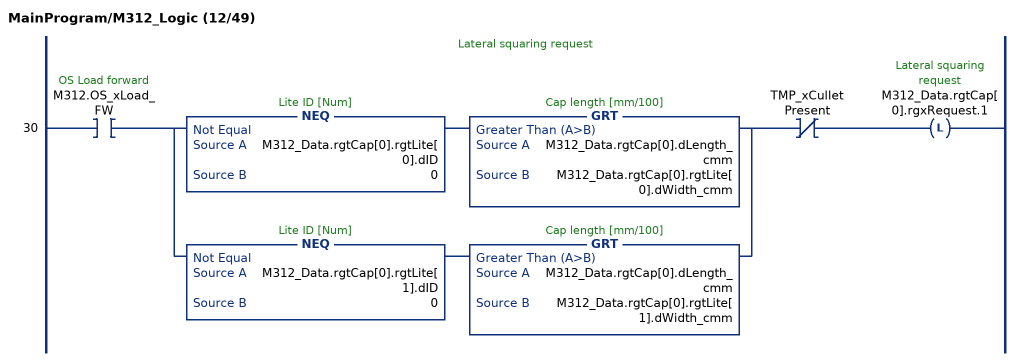
   // Lateral squaring request
   30: XIC(M312.OS_xLoad_FW)[NEQ(M312_Data.rgtCap[0].rgtLite[0].dID,0) GRT(M312_Data.rgtCap[0].dLength_cmm,M312_Data.rgtCap[0].rgtLite[0].dWidth_cmm) ,NEQ(M312_Data.rgtCap[0].rgtLite[1].dID,0) GRT(M312_Data.rgtCap[0].dLength_cmm,M312_Data.rgtCap[0].rgtLite[1].dWidth_cmm) ]XIO(TMP_xCulletPresent)OTL(M312_Data.rgtCap[0].rgxRequest.1);
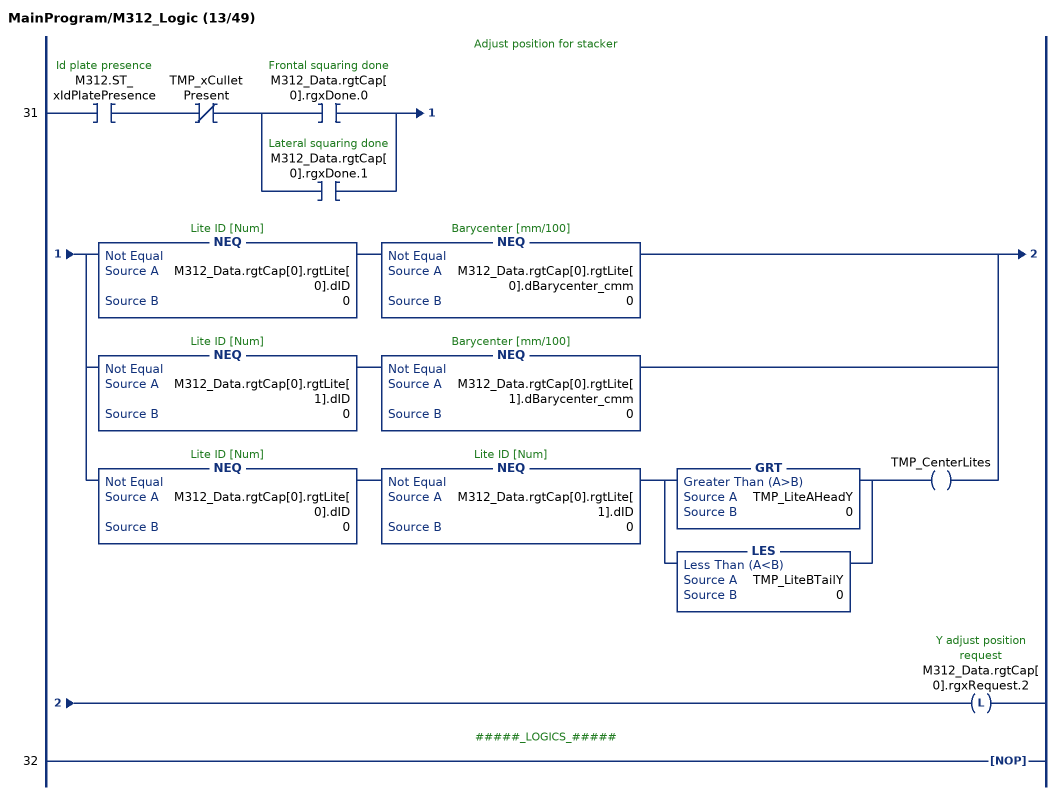
   // Adjust position for stacker
   31: XIC(M312.ST_xIdPlatePresence)XIO(TMP_xCulletPresent)[XIC(M312_Data.rgtCap[0].rgxDone.0) ,XIC(M312_Data.rgtCap[0].rgxDone.1) ][[NEQ(M312_Data.rgtCap[0].rgtLite[0].dID,0) NEQ(M312_Data.rgtCap[0].rgtLite[0].dBarycenter_cmm,0) ,NEQ(M312_Data.rgtCap[0].rgtLite[1].dID,0) NEQ(M312_Data.rgtCap[0].rgtLite[1].dBarycenter_cmm,0) ] ,NEQ(M312_Data.rgtCap[0].rgtLite[0].dID,0) NEQ(M312_Data.rgtCap[0].rgtLite[1].dID,0) [GRT(TMP_LiteAHeadY,0) ,LES(TMP_LiteBTailY,0) ] OTE(TMP_CenterLites) ]OTL(M312_Data.rgtCap[0].rgxRequest.2);
   // #####_LOGICS_#####
   32: NOP();
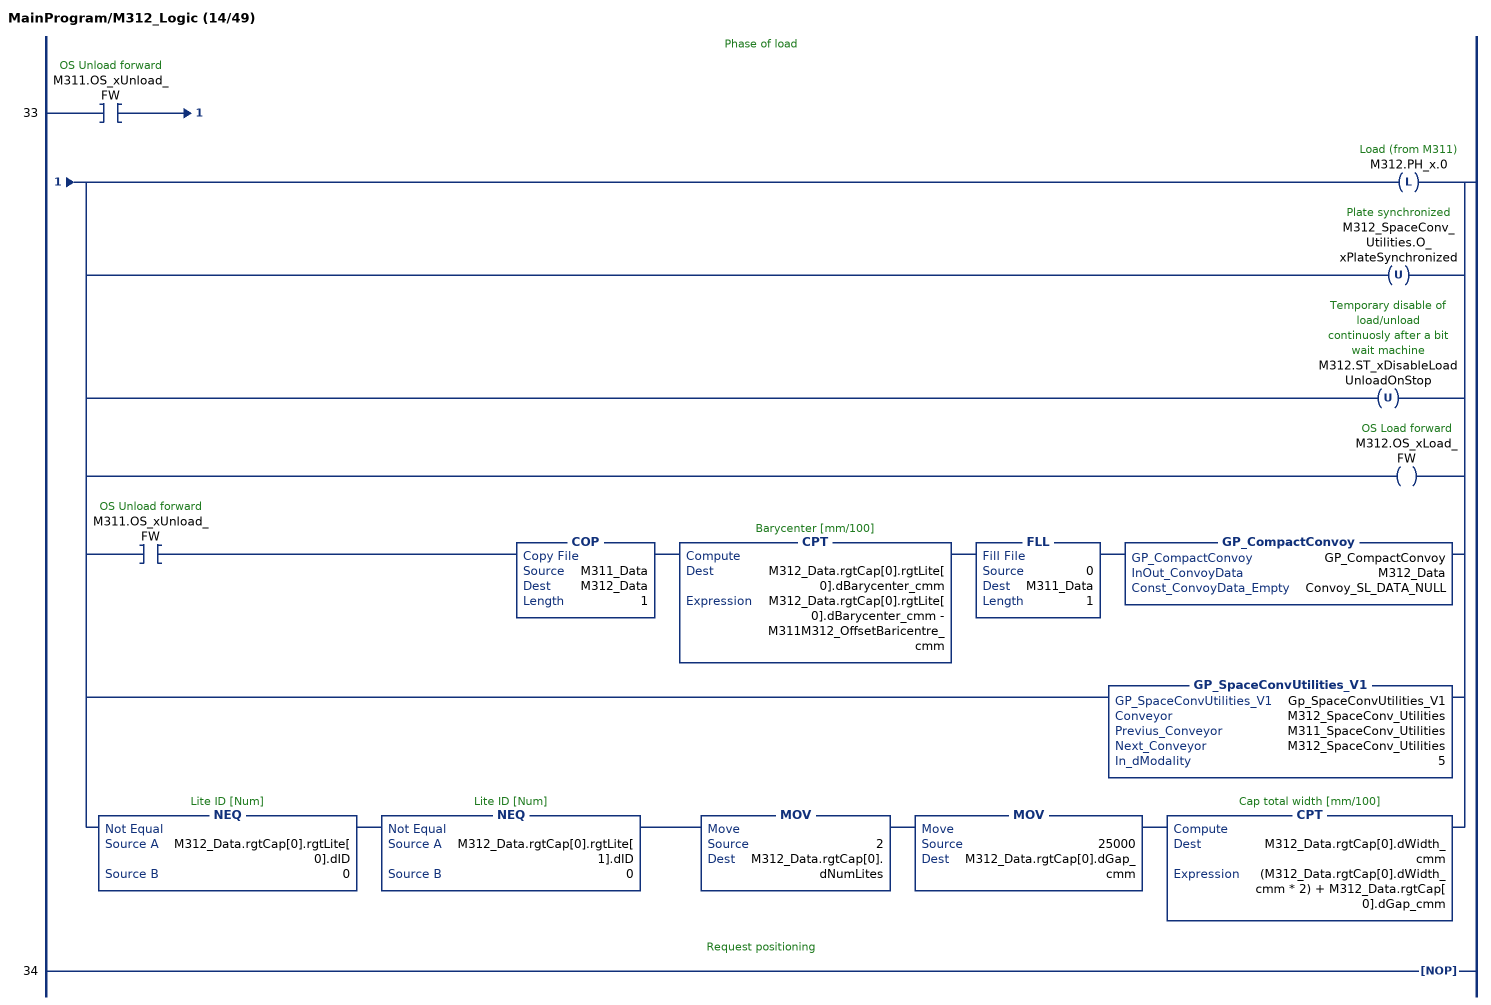
   // Phase of load
   33: XIC(M311.OS_xUnload_FW)[OTL(M312.PH_x.0) ,OTU(M312_SpaceConv_Utilities.O_xPlateSynchronized) ,OTU(M312.ST_xDisableLoadUnloadOnStop) ,OTE(M312.OS_xLoad_FW) ,XIC(M311.OS_xUnload_FW) COP(M311_Data,M312_Data,1) CPT(M312_Data.rgtCap[0].rgtLite[0].dBarycenter_cmm,M312_Data.rgtCap[0].rgtLite[0].dBarycenter_cmm - M311M312_OffsetBaricentre_cmm) FLL(0,M311_Data,1) GP_CompactConvoy(GP_CompactConvoy,M312_Data,Convoy_SL_DATA_NULL) ,GP_SpaceConvUtilities_V1(Gp_SpaceConvUtilities_V1,M312_SpaceConv_Utilities,M311_SpaceConv_Utilities,M312_SpaceConv_Utilities,5) ,NEQ(M312_Data.rgtCap[0].rgtLite[0].dID,0) NEQ(M312_Data.rgtCap[0].rgtLite[1].dID,0) MOV(2,M312_Data.rgtCap[0].dNumLites) MOV(25000,M312_Data.rgtCap[0].dGap_cmm) CPT(M312_Data.rgtCap[0].dWidth_cmm,(M312_Data.rgtCap[0].dWidth_cmm * 2) + M312_Data.rgtCap[0].dGap_cmm) ];
   // Request positioning
   34: NOP();
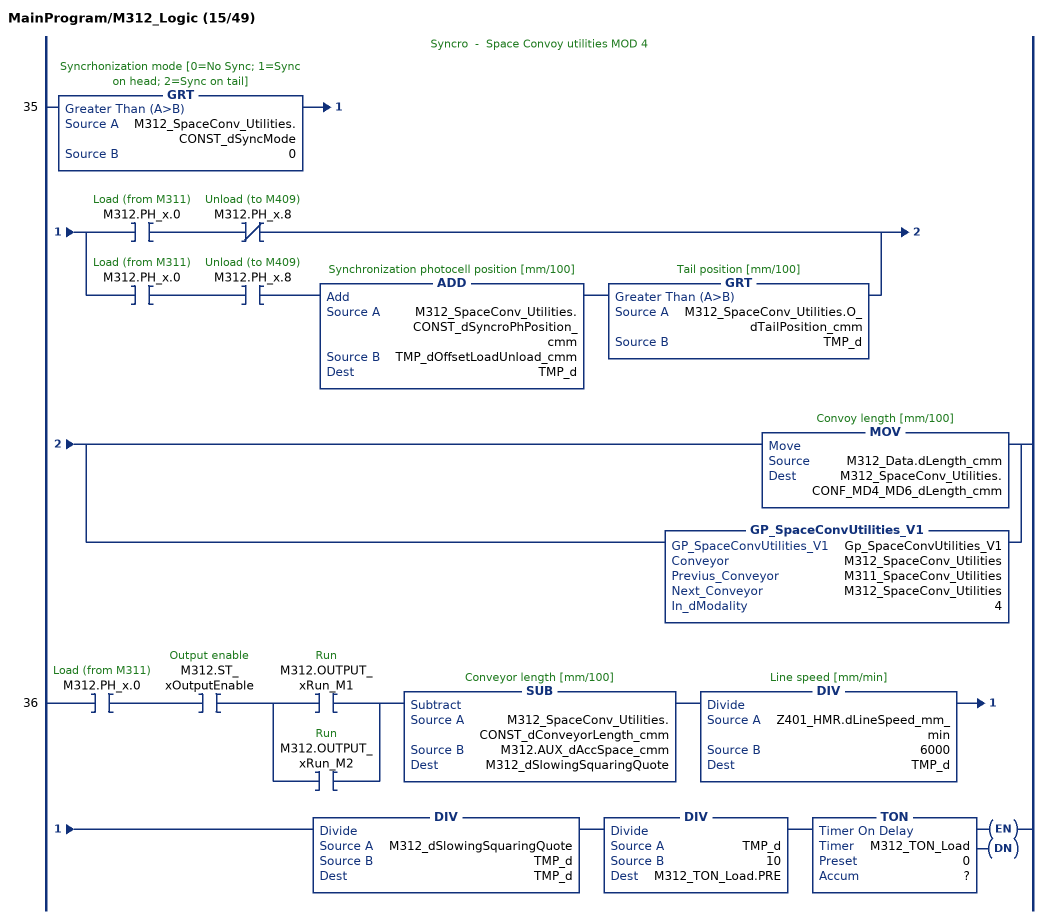
   // Syncro  -  Space Convoy utilities MOD 4
   35: GRT(M312_SpaceConv_Utilities.CONST_dSyncMode,0)[XIC(M312.PH_x.0) XIO(M312.PH_x.8) ,XIC(M312.PH_x.0) XIC(M312.PH_x.8) ADD(M312_SpaceConv_Utilities.CONST_dSyncroPhPosition_cmm,TMP_dOffsetLoadUnload_cmm,TMP_d) GRT(M312_SpaceConv_Utilities.O_dTailPosition_cmm,TMP_d) ][MOV(M312_Data.dLength_cmm,M312_SpaceConv_Utilities.CONF_MD4_MD6_dLength_cmm) ,GP_SpaceConvUtilities_V1(Gp_SpaceConvUtilities_V1,M312_SpaceConv_Utilities,M311_SpaceConv_Utilities,M312_SpaceConv_Utilities,4) ];
   36: XIC(M312.PH_x.0)XIC(M312.ST_xOutputEnable)[XIC(M312.OUTPUT_xRun_M1) ,XIC(M312.OUTPUT_xRun_M2) ]SUB(M312_SpaceConv_Utilities.CONST_dConveyorLength_cmm,M312.AUX_dAccSpace_cmm,M312_dSlowingSquaringQuote)DIV(Z401_HMR.dLineSpeed_mm_min,6000,TMP_d)DIV(M312_dSlowingSquaringQuote,TMP_d,TMP_d)DIV(TMP_d,10,M312_TON_Load.PRE)TON(M312_TON_Load,?,?);
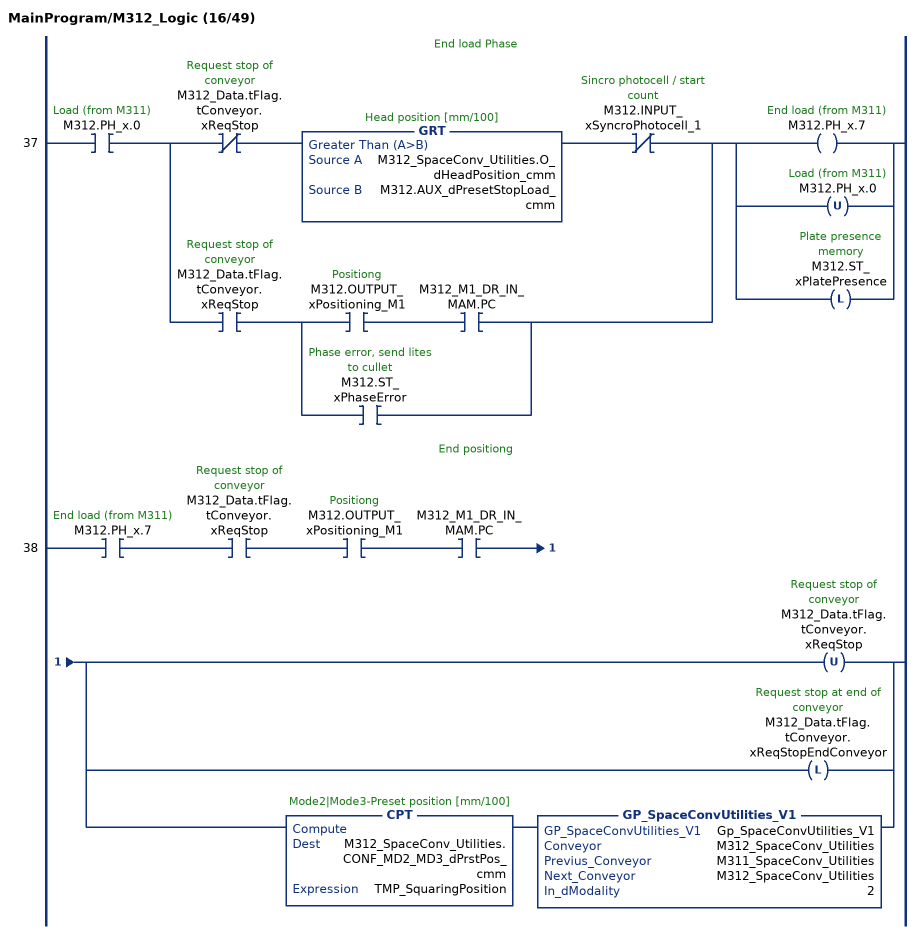
   // End load Phase
   37: XIC(M312.PH_x.0)[XIO(M312_Data.tFlag.tConveyor.xReqStop) GRT(M312_SpaceConv_Utilities.O_dHeadPosition_cmm,M312.AUX_dPresetStopLoad_cmm) XIO(M312.INPUT_xSyncroPhotocell_1) ,XIC(M312_Data.tFlag.tConveyor.xReqStop) [XIC(M312.OUTPUT_xPositioning_M1) XIC(M312_M1_DR_IN_MAM.PC) ,XIC(M312.ST_xPhaseError) ] ][OTE(M312.PH_x.7) ,OTU(M312.PH_x.0) ,OTL(M312.ST_xPlatePresence) ];
   // End positiong
   38: XIC(M312.PH_x.7)XIC(M312_Data.tFlag.tConveyor.xReqStop)XIC(M312.OUTPUT_xPositioning_M1)XIC(M312_M1_DR_IN_MAM.PC)[OTU(M312_Data.tFlag.tConveyor.xReqStop) ,OTL(M312_Data.tFlag.tConveyor.xReqStopEndConveyor) ,CPT(M312_SpaceConv_Utilities.CONF_MD2_MD3_dPrstPos_cmm,TMP_SquaringPosition) GP_SpaceConvUtilities_V1(Gp_SpaceConvUtilities_V1,M312_SpaceConv_Utilities,M311_SpaceConv_Utilities,M312_SpaceConv_Utilities,2) ];
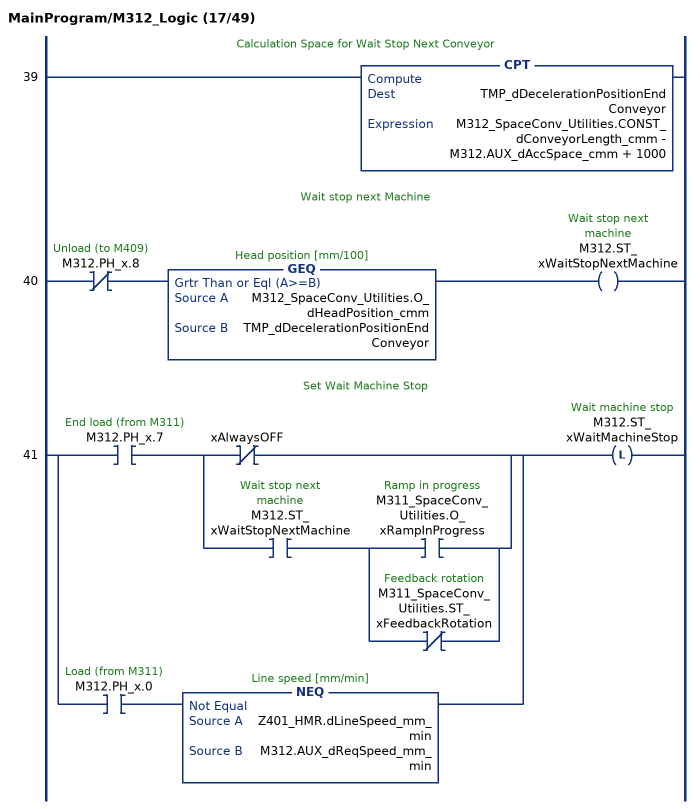
   // Calculation Space for Wait Stop Next Conveyor
   39: CPT(TMP_dDecelerationPositionEndConveyor,M312_SpaceConv_Utilities.CONST_dConveyorLength_cmm - M312.AUX_dAccSpace_cmm + 1000);
   // Wait stop next Machine
   40: XIO(M312.PH_x.8)GEQ(M312_SpaceConv_Utilities.O_dHeadPosition_cmm,TMP_dDecelerationPositionEndConveyor)OTE(M312.ST_xWaitStopNextMachine);
   // Set Wait Machine Stop
   41: [XIC(M312.PH_x.7) [XIO(xAlwaysOFF) ,XIC(M312.ST_xWaitStopNextMachine) [XIC(M311_SpaceConv_Utilities.O_xRampInProgress) ,XIO(M311_SpaceConv_Utilities.ST_xFeedbackRotation) ] ] ,XIC(M312.PH_x.0) NEQ(Z401_HMR.dLineSpeed_mm_min,M312.AUX_dReqSpeed_mm_min) ]OTL(M312.ST_xWaitMachineStop);
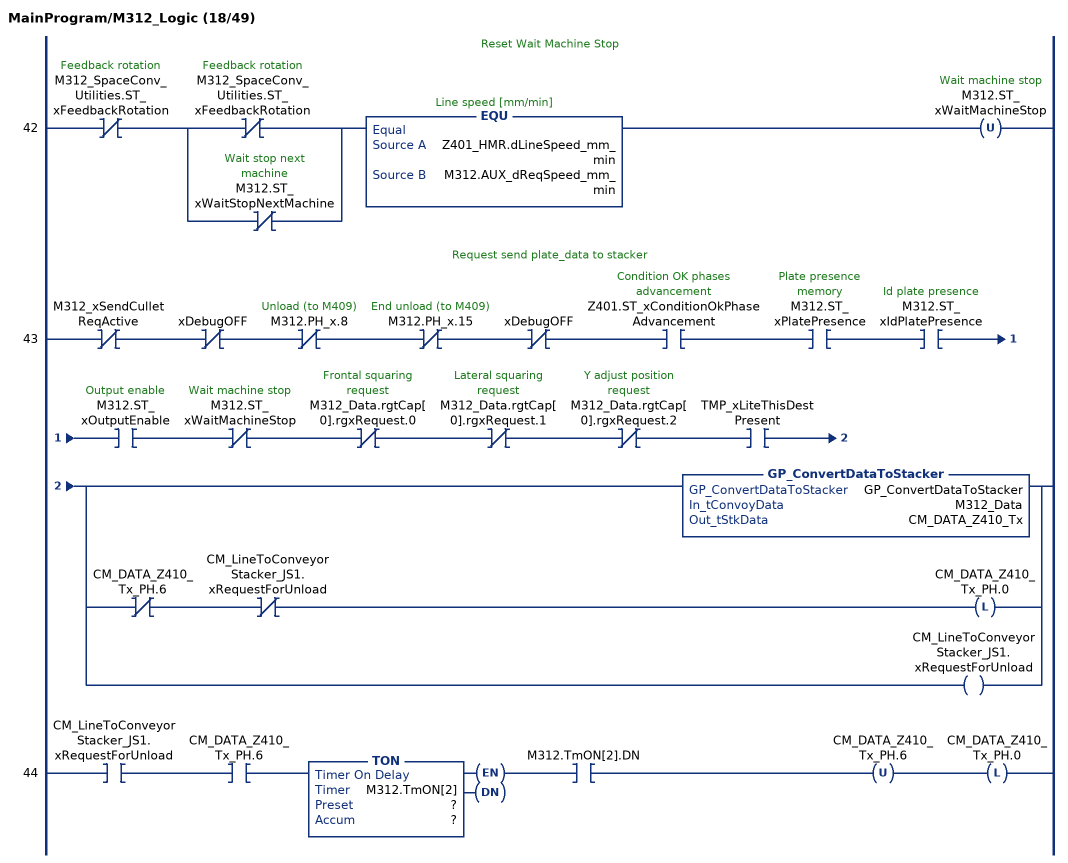
   // Reset Wait Machine Stop
   42: XIO(M312_SpaceConv_Utilities.ST_xFeedbackRotation)[XIO(M312_SpaceConv_Utilities.ST_xFeedbackRotation) ,XIO(M312.ST_xWaitStopNextMachine) ]EQU(Z401_HMR.dLineSpeed_mm_min,M312.AUX_dReqSpeed_mm_min)OTU(M312.ST_xWaitMachineStop);
   // Request send plate_data to stacker
   43: XIO(M312_xSendCulletReqActive)XIO(xDebugOFF)XIO(M312.PH_x.8)XIO(M312.PH_x.15)XIO(xDebugOFF)XIC(Z401.ST_xConditionOkPhaseAdvancement)XIC(M312.ST_xPlatePresence)XIC(M312.ST_xIdPlatePresence)XIC(M312.ST_xOutputEnable)XIO(M312.ST_xWaitMachineStop)XIO(M312_Data.rgtCap[0].rgxRequest.0)XIO(M312_Data.rgtCap[0].rgxRequest.1)XIO(M312_Data.rgtCap[0].rgxRequest.2)XIC(TMP_xLiteThisDestPresent)[GP_ConvertDataToStacker(GP_ConvertDataToStacker,M312_Data,CM_DATA_Z410_Tx) ,XIO(CM_DATA_Z410_Tx_PH.6) XIO(CM_LineToConveyorStacker_JS1.xRequestForUnload) OTL(CM_DATA_Z410_Tx_PH.0) ,OTE(CM_LineToConveyorStacker_JS1.xRequestForUnload) ];
   44: XIC(CM_LineToConveyorStacker_JS1.xRequestForUnload)XIC(CM_DATA_Z410_Tx_PH.6)TON(M312.TmON[2],?,?)XIC(M312.TmON[2].DN)OTU(CM_DATA_Z410_Tx_PH.6)OTL(CM_DATA_Z410_Tx_PH.0);
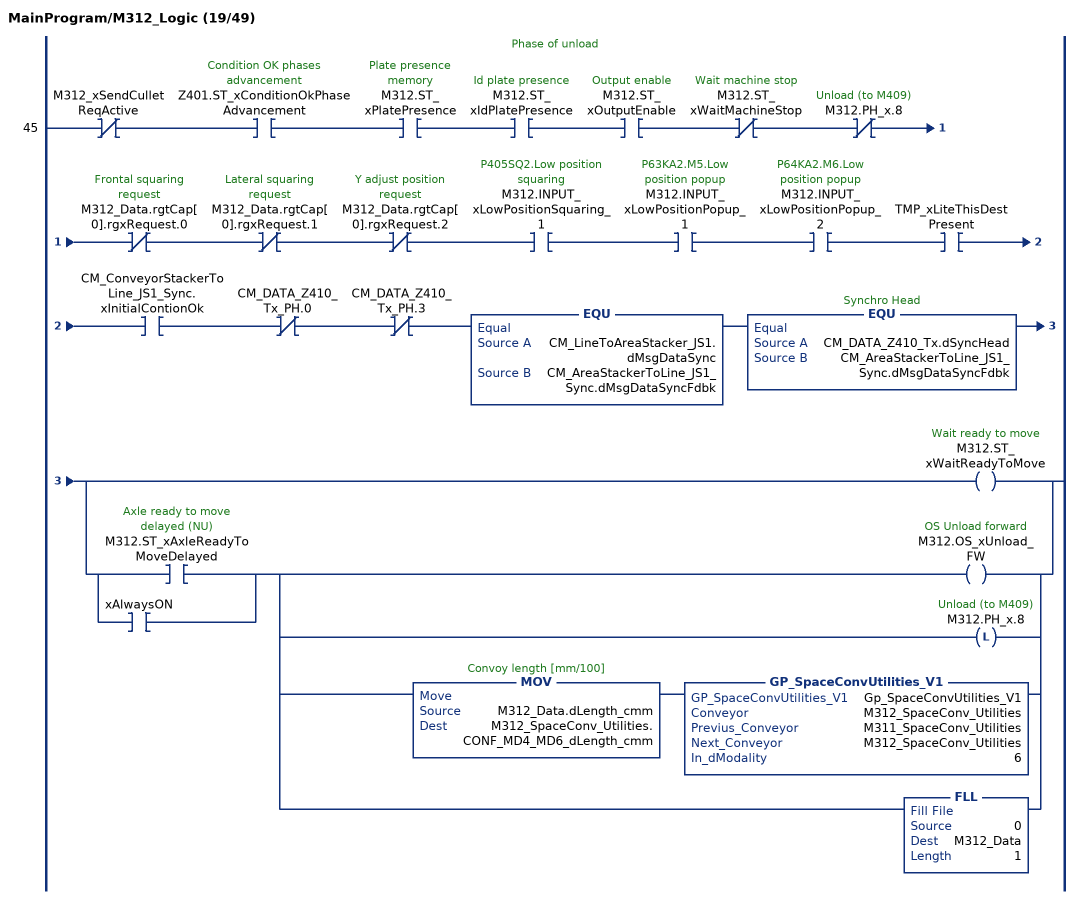
   // Phase of unload
   45: XIO(M312_xSendCulletReqActive)XIC(Z401.ST_xConditionOkPhaseAdvancement)XIC(M312.ST_xPlatePresence)XIC(M312.ST_xIdPlatePresence)XIC(M312.ST_xOutputEnable)XIO(M312.ST_xWaitMachineStop)XIO(M312.PH_x.8)XIO(M312_Data.rgtCap[0].rgxRequest.0)XIO(M312_Data.rgtCap[0].rgxRequest.1)XIO(M312_Data.rgtCap[0].rgxRequest.2)XIC(M312.INPUT_xLowPositionSquaring_1)XIC(M312.INPUT_xLowPositionPopup_1)XIC(M312.INPUT_xLowPositionPopup_2)XIC(TMP_xLiteThisDestPresent)XIC(CM_ConveyorStackerToLine_JS1_Sync.xInitialContionOk)XIO(CM_DATA_Z410_Tx_PH.0)XIO(CM_DATA_Z410_Tx_PH.3)EQU(CM_LineToAreaStacker_JS1.dMsgDataSync,CM_AreaStackerToLine_JS1_Sync.dMsgDataSyncFdbk)EQU(CM_DATA_Z410_Tx.dSyncHead,CM_AreaStackerToLine_JS1_Sync.dMsgDataSyncFdbk)[OTE(M312.ST_xWaitReadyToMove) ,[XIC(M312.ST_xAxleReadyToMoveDelayed) ,XIC(xAlwaysON) ] [OTE(M312.OS_xUnload_FW) ,OTL(M312.PH_x.8) ,MOV(M312_Data.dLength_cmm,M312_SpaceConv_Utilities.CONF_MD4_MD6_dLength_cmm) GP_SpaceConvUtilities_V1(Gp_SpaceConvUtilities_V1,M312_SpaceConv_Utilities,M311_SpaceConv_Utilities,M312_SpaceConv_Utilities,6) ,FLL(0,M312_Data,1) ] ];
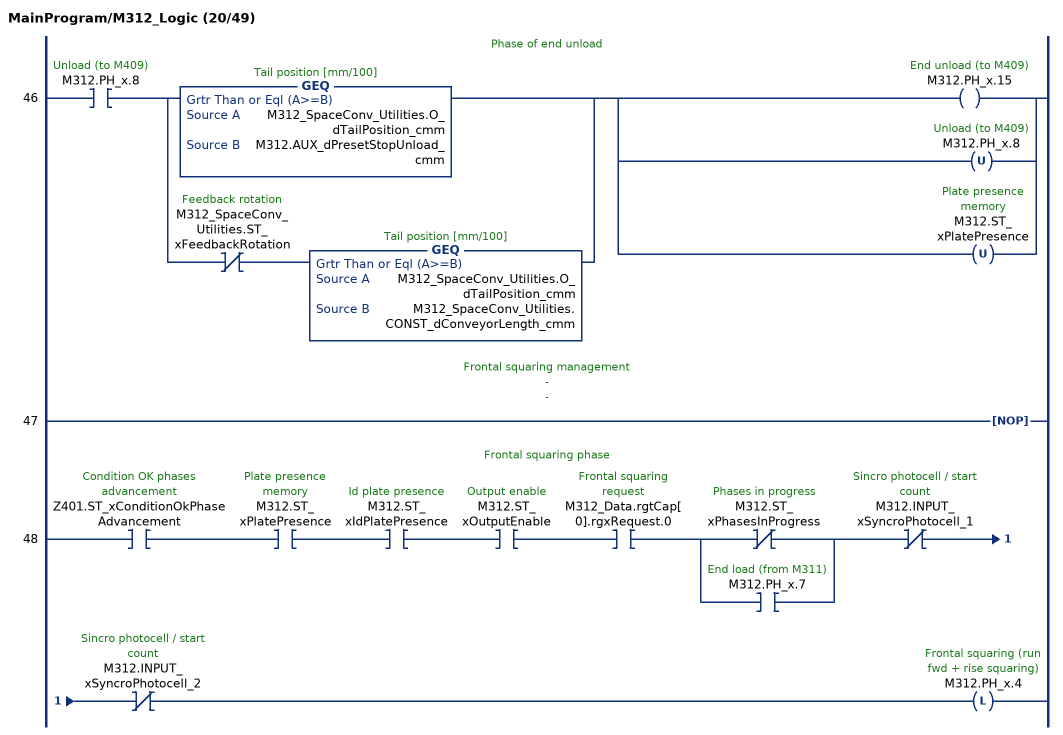
   // Phase of end unload
   46: XIC(M312.PH_x.8)[GEQ(M312_SpaceConv_Utilities.O_dTailPosition_cmm,M312.AUX_dPresetStopUnload_cmm) ,XIO(M312_SpaceConv_Utilities.ST_xFeedbackRotation) GEQ(M312_SpaceConv_Utilities.O_dTailPosition_cmm,M312_SpaceConv_Utilities.CONST_dConveyorLength_cmm) ][OTE(M312.PH_x.15) ,OTU(M312.PH_x.8) ,OTU(M312.ST_xPlatePresence) ];
   // Frontal squaring management
   // -
   // -
   47: NOP();
   // Frontal squaring phase
   48: XIC(Z401.ST_xConditionOkPhaseAdvancement)XIC(M312.ST_xPlatePresence)XIC(M312.ST_xIdPlatePresence)XIC(M312.ST_xOutputEnable)XIC(M312_Data.rgtCap[0].rgxRequest.0)[XIO(M312.ST_xPhasesInProgress) ,XIC(M312.PH_x.7) ]XIO(M312.INPUT_xSyncroPhotocell_1)XIO(M312.INPUT_xSyncroPhotocell_2)OTL(M312.PH_x.4);
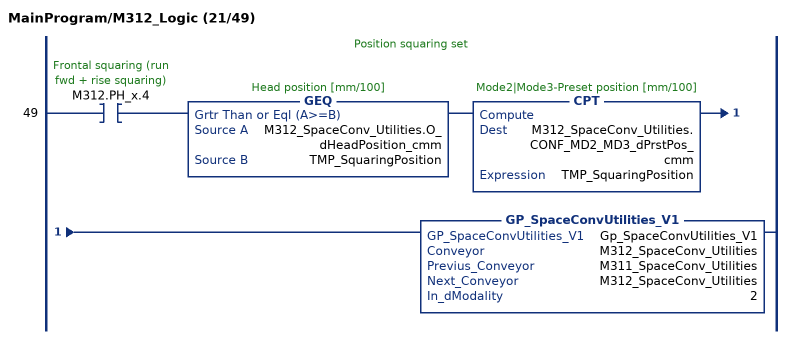
   // Position squaring set
   49: XIC(M312.PH_x.4)GEQ(M312_SpaceConv_Utilities.O_dHeadPosition_cmm,TMP_SquaringPosition)CPT(M312_SpaceConv_Utilities.CONF_MD2_MD3_dPrstPos_cmm,TMP_SquaringPosition)GP_SpaceConvUtilities_V1(Gp_SpaceConvUtilities_V1,M312_SpaceConv_Utilities,M311_SpaceConv_Utilities,M312_SpaceConv_Utilities,2);
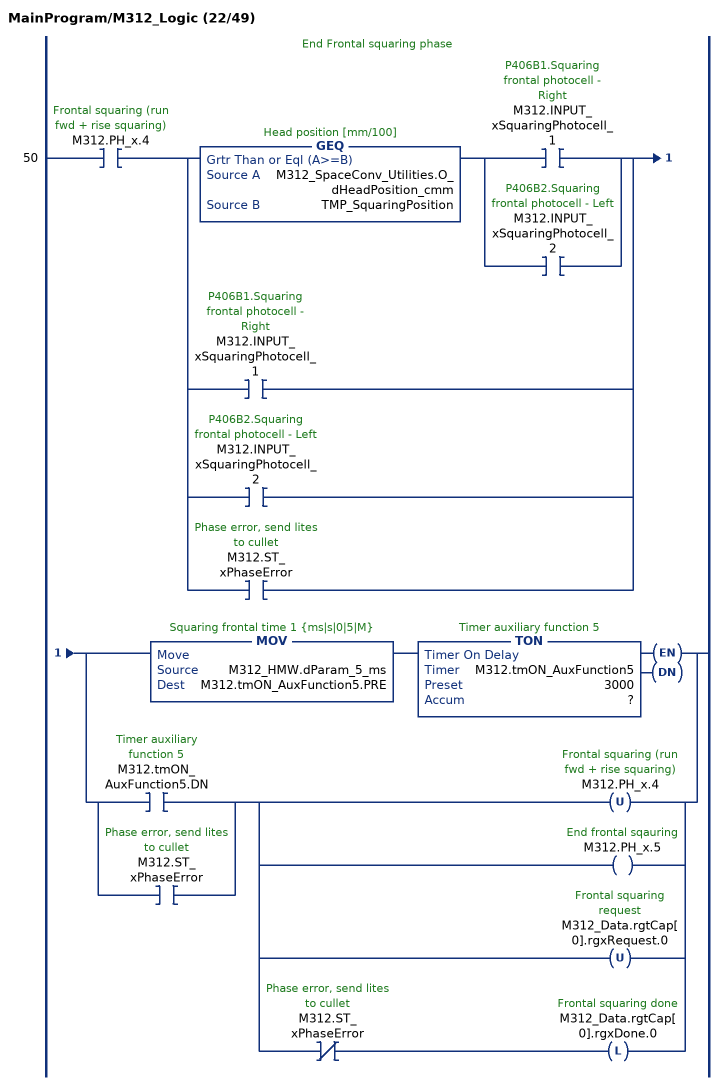
   // End Frontal squaring phase
   50: XIC(M312.PH_x.4)[[GEQ(M312_SpaceConv_Utilities.O_dHeadPosition_cmm,TMP_SquaringPosition) [XIC(M312.INPUT_xSquaringPhotocell_1) ,XIC(M312.INPUT_xSquaringPhotocell_2) ] ,XIC(M312.INPUT_xSquaringPhotocell_1) ,XIC(M312.INPUT_xSquaringPhotocell_2) ] ,XIC(M312.ST_xPhaseError) ][MOV(M312_HMW.dParam_5_ms,M312.tmON_AuxFunction5.PRE) TON(M312.tmON_AuxFunction5,?,?) ,[XIC(M312.tmON_AuxFunction5.DN) ,XIC(M312.ST_xPhaseError) ] [OTU(M312.PH_x.4) ,OTE(M312.PH_x.5) ,OTU(M312_Data.rgtCap[0].rgxRequest.0) ,XIO(M312.ST_xPhaseError) OTL(M312_Data.rgtCap[0].rgxDone.0) ] ];
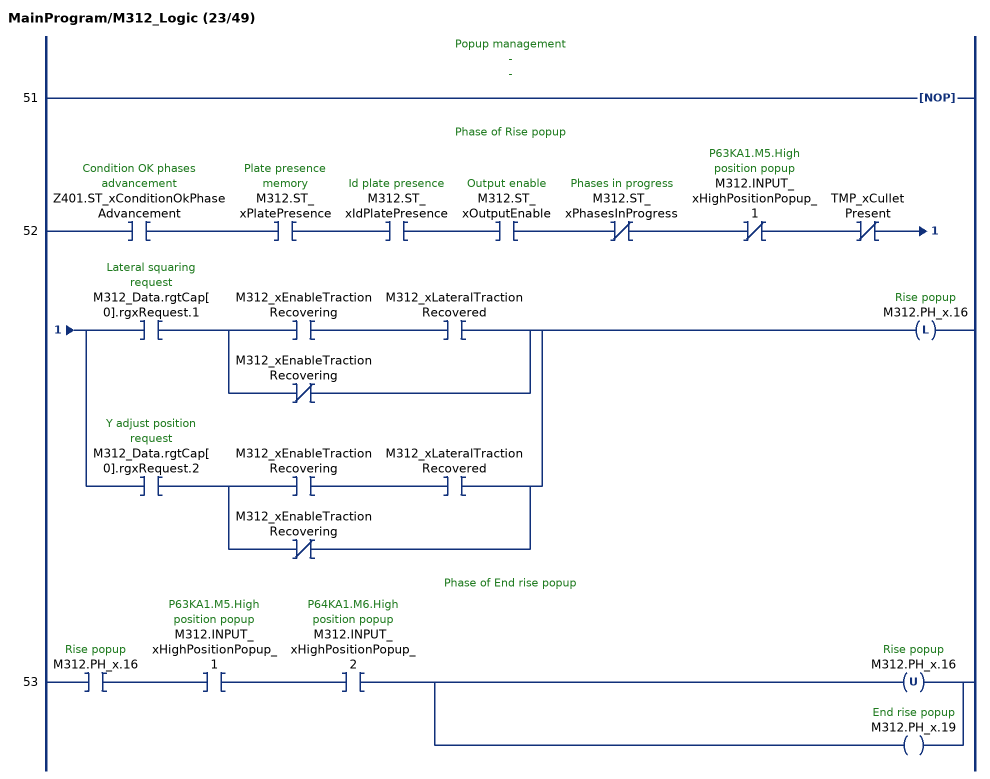
   // Popup management
   // -
   // -
   51: NOP();
   // Phase of Rise popup
   52: XIC(Z401.ST_xConditionOkPhaseAdvancement)XIC(M312.ST_xPlatePresence)XIC(M312.ST_xIdPlatePresence)XIC(M312.ST_xOutputEnable)XIO(M312.ST_xPhasesInProgress)XIO(M312.INPUT_xHighPositionPopup_1)XIO(TMP_xCulletPresent)[XIC(M312_Data.rgtCap[0].rgxRequest.1) [XIC(M312_xEnableTractionRecovering) XIC(M312_xLateralTractionRecovered) ,XIO(M312_xEnableTractionRecovering) ] ,XIC(M312_Data.rgtCap[0].rgxRequest.2) [XIC(M312_xEnableTractionRecovering) XIC(M312_xLateralTractionRecovered) ,XIO(M312_xEnableTractionRecovering) ] ]OTL(M312.PH_x.16);
   // Phase of End rise popup
   53: XIC(M312.PH_x.16)XIC(M312.INPUT_xHighPositionPopup_1)XIC(M312.INPUT_xHighPositionPopup_2)[OTU(M312.PH_x.16) ,OTE(M312.PH_x.19) ];
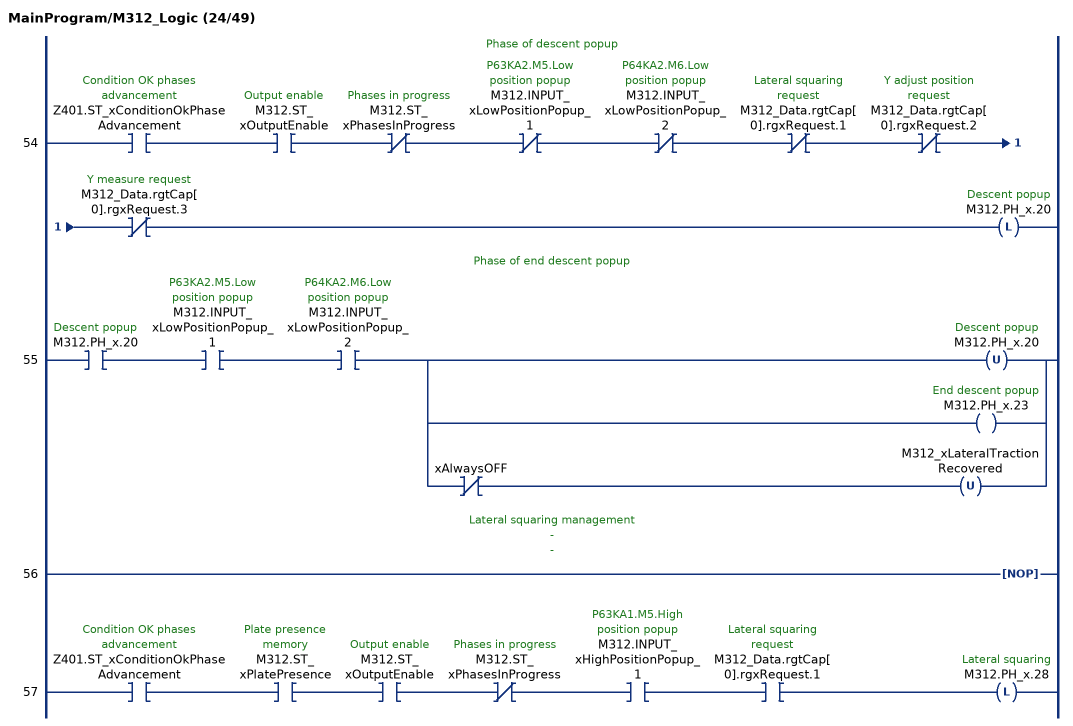
   // Phase of descent popup
   54: XIC(Z401.ST_xConditionOkPhaseAdvancement)XIC(M312.ST_xOutputEnable)XIO(M312.ST_xPhasesInProgress)XIO(M312.INPUT_xLowPositionPopup_1)XIO(M312.INPUT_xLowPositionPopup_2)XIO(M312_Data.rgtCap[0].rgxRequest.1)XIO(M312_Data.rgtCap[0].rgxRequest.2)XIO(M312_Data.rgtCap[0].rgxRequest.3)OTL(M312.PH_x.20);
   // Phase of end descent popup
   55: XIC(M312.PH_x.20)XIC(M312.INPUT_xLowPositionPopup_1)XIC(M312.INPUT_xLowPositionPopup_2)[OTU(M312.PH_x.20) ,OTE(M312.PH_x.23) ,XIO(xAlwaysOFF) OTU(M312_xLateralTractionRecovered) ];
   // Lateral squaring management
   // -
   // -
   56: NOP();
   57: XIC(Z401.ST_xConditionOkPhaseAdvancement)XIC(M312.ST_xPlatePresence)XIC(M312.ST_xOutputEnable)XIO(M312.ST_xPhasesInProgress)XIC(M312.INPUT_xHighPositionPopup_1)XIC(M312_Data.rgtCap[0].rgxRequest.1)OTL(M312.PH_x.28);
